(* Logix 5000 project; controller FV vendor 1 type 14 code 217 rev 31.11; software revision 31.00; part 63 of 63 *)
(* tags used below, declared in another part *)
   Alarm_Reset : BOOL;
   CWD : CHECKWORD_FLAGS;
   Default_Check_Time : DINT;
   Item_Faults_Are_Latched : BOOL;
   Item_Simulation_Flag : BOOL;
   One_Second_One_Scan : ALIAS FOR One_Second_1_scan;
   YP_AV1 : PlantItem;   // AV1
   YP_AV1_ALARM : ALARM_DIGITAL;
   YP_AV1_DR : ALIAS FOR RIO_Rack_3:3:O.Data.3;
   YP_AV1_O : ALIAS FOR RIO_Rack_3:1:I.Data.0;
   YP_AV2 : PlantItem;   // AV2
   YP_AV2_ALARM : ALARM_DIGITAL;
   YP_AV2_DR : ALIAS FOR RIO_Rack_3:3:O.Data.5;
   YP_AV2_O : ALIAS FOR RIO_Rack_3:1:I.Data.2;
   YP_AV3 : PlantItem;   // AV3
   YP_AV3_ALARM : ALARM_DIGITAL;
   YP_AV3_DR : ALIAS FOR RIO_Rack_3:3:O.Data.6;
   YP_AV3_O : ALIAS FOR RIO_Rack_3:1:I.Data.4;
   YP_AV4 : PlantItem;   // AV4
   YP_AV4_ALARM : ALARM_DIGITAL;
   YP_AV4_DR : ALIAS FOR RIO_Rack_3:3:O.Data.7;
   YP_AV4_O : ALIAS FOR RIO_Rack_3:1:I.Data.6;
   YP_AV5 : PlantItem;   // AV5
   YP_AV5_ALARM : ALARM_DIGITAL;
   YP_AV5_DR : ALIAS FOR RIO_Rack_3:3:O.Data.8;
   YP_AV5_O : ALIAS FOR RIO_Rack_3:1:I.Data.8;
   YP_AV6 : PlantItem;   // AV6
   YP_AV6_ALARM : ALARM_DIGITAL;
   YP_AV6_DR : ALIAS FOR RIO_Rack_3:3:O.Data.9;
   YP_AV6_O : ALIAS FOR RIO_Rack_3:1:I.Data.10;
   YP_AV7 : PlantItem;   // AV7
   YP_AV7_ALARM : ALARM_DIGITAL;
   YP_AV7_DR : ALIAS FOR RIO_Rack_3:3:O.Data.10;
   YP_AV7_O : ALIAS FOR RIO_Rack_3:1:I.Data.12;
   YP_AV8 : PlantItem;   // AV8
   YP_AV8_ALARM : ALARM_DIGITAL;
   YP_AV8_DR : ALIAS FOR RIO_Rack_3:3:O.Data.11;
   YP_AV8_O : ALIAS FOR RIO_Rack_3:1:I.Data.14;
   YP_B103 : INT[15];   // Original N File From SLC, No Description Available
   YP_B3 : INT[7];   // BINARY
   YP_B30 : INT[37];   // Original N File From SLC, No Description Available
   YP_N40 : INT[9];   // Original N File From SLC, No Description Available
   YP_N50 : INT[15];   // Original N File From SLC, No Description Available
   YP_N55 : INT[244];   // Original N File From SLC, No Description Available
   YP_N7 : INT[56];   // INTEGER
   YP_T4 : TIMER[16];   // TIMER
   YP_YST1_HL : PlantItem;   // YST1_HL
   YP_YST2_HL : PlantItem;   // YST2_HL
(* YP_Common, continued *)

ROUTINE YP_RQD_FLAGS_17   (* ladder *)
   0: [XIC(YP_N40[0].1) ,XIC(YP_N40[1].1) ]OTE(YP_B30[0].1);
   1: [XIC(YP_N40[0].3) ,XIC(YP_N40[0].4) ]XIC(YP_B3[0].10)XIC(YP_B3[0].8)[XIC(YP_B3[0].0) ,XIC(YP_B3[0].2) ,XIC(YP_B3[0].4) ,XIC(YP_B3[0].6) ]OTE(YP_B30[0].4);
   2: [[XIC(YP_N40[0].3) ,XIC(YP_N40[0].4) ,XIC(YP_B103[2].0) ] EQU(YP_N50[5],0) ,EQU(YP_N50[5],1) ]OTE(YP_B30[0].9);
   3: [[XIC(YP_N40[0].3) ,XIC(YP_N40[0].4) ,XIC(YP_B103[2].1) ] EQU(YP_N50[4],0) ,EQU(YP_N50[4],1) ]OTE(YP_B30[0].8);
   4: [[XIC(YP_N40[0].3) ,XIC(YP_N40[0].4) ,XIC(YP_B103[2].0) ,XIC(YP_B103[2].1) ] EQU(YP_N50[0],0) ,EQU(YP_N50[0],1) ]OTE(YP_B30[0].3);
   5: [[XIC(YP_N40[0].3) ,XIC(YP_N40[0].4) ,XIC(YP_B103[2].0) ] EQU(YP_N50[1],0) ,EQU(YP_N50[1],1) ]OTE(YP_B30[0].5);
   6: [[XIC(YP_N40[0].4) ,XIC(YP_B103[2].0) ] EQU(YP_N50[2],0) ,EQU(YP_N50[2],1) ]OTE(YP_B30[0].6);
   7: [[XIC(YP_N40[0].4) ,XIC(YP_B103[2].0) ] EQU(YP_N50[3],0) ,EQU(YP_N50[3],1) ]OTE(YP_B30[0].7);
   8: [XIC(YP_N40[0].7) ,XIC(YP_N40[1].5) ]OTE(YP_B30[0].0);
   9: XIC(YP_N40[0].8)OTE(YP_B30[0].2);
   10: [XIC(YP_N40[2].1) EQU(YP_N50[7],0) ,EQU(YP_N50[7],1) ]OTE(YP_B30[0].11);
   11: [XIC(YP_N40[3].1) EQU(YP_N50[6],0) XIO(YP_N7[38].0) XIO(YP_N7[38].1) ,EQU(YP_N50[6],1) ]OTE(YP_B30[0].10);
   12: [[XIC(YP_N40[0].3) ,XIC(YP_N40[0].4) ] XIC(YP_B3[0].10) XIC(YP_B3[0].8) [XIC(YP_B3[0].0) ,XIC(YP_B3[0].2) ,XIC(YP_B3[0].4) ,XIC(YP_B3[0].6) ] EQU(YP_N50[8],0) ,EQU(YP_N50[8],1) ]OTE(YP_B30[0].12);
   13: [XIC(YP_N40[3].1) XIC(YP_B3[0].12) EQU(YP_N50[9],0) ,EQU(YP_N50[9],1) ]OTE(YP_B30[0].14);
   14: XIC(YP_N40[0].0)MOV(0,YP_N55[2]);
   15: [XIC(YP_N40[0].1) ,XIC(YP_N40[1].1) ]MOV(1,YP_N55[2]);
   16: [XIC(YP_N40[0].2) ,XIC(YP_N40[1].2) ]MOV(2,YP_N55[2]);
   17: XIC(YP_N40[0].3)MOV(3,YP_N55[2]);
   18: XIC(YP_N40[0].4)MOV(4,YP_N55[2]);
   19: XIC(YP_N40[0].5)MOV(5,YP_N55[2]);
   20: XIC(YP_N40[0].6)MOV(6,YP_N55[2]);
   21: [XIC(YP_N40[0].7) ,XIC(YP_N40[1].5) ]MOV(7,YP_N55[2]);
   22: XIC(YP_N40[0].8)MOV(8,YP_N55[2]);
   23: EQU(YP_N55[0],1)MOV(9,YP_N55[2]);
   24: XIC(YP_N40[1].2)MOV(10,YP_N55[2]);
   25: XIC(YP_N40[1].3)MOV(11,YP_N55[2]);
   26: XIC(YP_N40[1].4)MOV(12,YP_N55[2]);
END_ROUTINE

ROUTINE YP_Valves   (* ladder *)
   0: [NEQ(YP_AV1.DriveBits,0) OTE(YP_AV1.CW.[CWD.AUTODRV]) ,[XIC(YP_AV1.CW.[CWD.AUTODRV]) XIO(YP_AV1.CW.[CWD.MANUAL]) ,XIC(YP_AV1.CW.[CWD.MANDRV]) XIC(YP_AV1.CW.[CWD.MANUAL]) ] OTE(YP_AV1.CW.[CWD.OUTPUT]) ,XIC(YP_AV1.CW.[CWD.OUTPUT]) OTE(YP_AV1_DR) ,XIC(S:FS) [OTU(YP_AV1.CW.[CWD.MANUAL]) ,LEQ(YP_AV1.CheckTime,0) MOV(Default_Check_Time,YP_AV1.CheckTime) ] ,[[XIC(YP_AV1_O) XIO(Item_Simulation_Flag) ,XIC(Item_Simulation_Flag) XIC(YP_AV1.CW.[CWD.OUTPUT]) XIO(YP_AV1.CW.[CWD.SIMFAIL]) ] OTE(YP_AV1.CW.[CWD.OPENFB]) ,[XIO(YP_AV1_O) XIO(Item_Simulation_Flag) ,XIC(Item_Simulation_Flag) XIO(YP_AV1.CW.[CWD.OUTPUT]) XIO(YP_AV1.CW.[CWD.SIMFAIL]) ] OTE(YP_AV1.CW.[CWD.CLOSEDFB]) ] ,[XIC(YP_AV1.CW.[CWD.OUTPUT]) XIO(YP_AV1.CW.[CWD.PREVSCAN]) ,XIO(YP_AV1.CW.[CWD.OUTPUT]) XIC(YP_AV1.CW.[CWD.PREVSCAN]) ] CLR(YP_AV1.CheckTimer) ,XIC(One_Second_One_Scan) LES(YP_AV1.CheckTimer,YP_AV1.CheckTime) ADD(YP_AV1.CheckTimer,1,YP_AV1.CheckTimer) ,XIO(YP_AV1.CW.[CWD.FAULT]) OTU(YP_AV1.CW.[CWD.FAULTLOGGED]) ,[GEQ(YP_AV1.CheckTimer,YP_AV1.CheckTime) [XIC(YP_AV1.CW.[CWD.OUTPUT]) [XIO(YP_AV1.CW.[CWD.OPENFB]) ,XIC(YP_AV1.CW.[CWD.CLOSEDFB]) ] ,XIO(YP_AV1.CW.[CWD.OUTPUT]) [XIC(YP_AV1.CW.[CWD.OPENFB]) ,XIO(YP_AV1.CW.[CWD.CLOSEDFB]) ] ] ,XIC(YP_AV1.CW.[CWD.FAULT]) XIC(Item_Faults_Are_Latched) ,XIC(YP_AV1.CW.[CWD.HIGHLIGHT]) ] XIO(YP_AV1.CW.[CWD.CHECKOFF]) XIO(Alarm_Reset) [OTE(YP_AV1.CW.[CWD.FAULT]) ,ALMD(YP_AV1_ALARM,0,0,0,0) ] ,XIC(YP_AV1.CW.[CWD.OUTPUT]) OTE(YP_AV1.CW.[CWD.PREVSCAN]) ];
   1: [NEQ(YP_AV2.DriveBits,0) OTE(YP_AV2.CW.[CWD.AUTODRV]) ,[XIC(YP_AV2.CW.[CWD.AUTODRV]) XIO(YP_AV2.CW.[CWD.MANUAL]) ,XIC(YP_AV2.CW.[CWD.MANDRV]) XIC(YP_AV2.CW.[CWD.MANUAL]) ] OTE(YP_AV2.CW.[CWD.OUTPUT]) ,XIC(YP_AV2.CW.[CWD.OUTPUT]) OTE(YP_AV2_DR) ,XIC(S:FS) [OTU(YP_AV2.CW.[CWD.MANUAL]) ,LEQ(YP_AV2.CheckTime,0) MOV(Default_Check_Time,YP_AV2.CheckTime) ] ,[[XIC(YP_AV2_O) XIO(Item_Simulation_Flag) ,XIC(Item_Simulation_Flag) XIC(YP_AV2.CW.[CWD.OUTPUT]) XIO(YP_AV2.CW.[CWD.SIMFAIL]) ] OTE(YP_AV2.CW.[CWD.OPENFB]) ,[XIO(YP_AV2_O) XIO(Item_Simulation_Flag) ,XIC(Item_Simulation_Flag) XIO(YP_AV2.CW.[CWD.OUTPUT]) XIO(YP_AV2.CW.[CWD.SIMFAIL]) ] OTE(YP_AV2.CW.[CWD.CLOSEDFB]) ] ,[XIC(YP_AV2.CW.[CWD.OUTPUT]) XIO(YP_AV2.CW.[CWD.PREVSCAN]) ,XIO(YP_AV2.CW.[CWD.OUTPUT]) XIC(YP_AV2.CW.[CWD.PREVSCAN]) ] CLR(YP_AV2.CheckTimer) ,XIC(One_Second_One_Scan) LES(YP_AV2.CheckTimer,YP_AV2.CheckTime) ADD(YP_AV2.CheckTimer,1,YP_AV2.CheckTimer) ,XIO(YP_AV2.CW.[CWD.FAULT]) OTU(YP_AV2.CW.[CWD.FAULTLOGGED]) ,[GEQ(YP_AV2.CheckTimer,YP_AV2.CheckTime) [XIC(YP_AV2.CW.[CWD.OUTPUT]) [XIO(YP_AV2.CW.[CWD.OPENFB]) ,XIC(YP_AV2.CW.[CWD.CLOSEDFB]) ] ,XIO(YP_AV2.CW.[CWD.OUTPUT]) [XIC(YP_AV2.CW.[CWD.OPENFB]) ,XIO(YP_AV2.CW.[CWD.CLOSEDFB]) ] ] ,XIC(YP_AV2.CW.[CWD.FAULT]) XIC(Item_Faults_Are_Latched) ,XIC(YP_AV2.CW.[CWD.HIGHLIGHT]) ] XIO(YP_AV2.CW.[CWD.CHECKOFF]) XIO(Alarm_Reset) [OTE(YP_AV2.CW.[CWD.FAULT]) ,ALMD(YP_AV2_ALARM,0,0,0,0) ] ,XIC(YP_AV2.CW.[CWD.OUTPUT]) OTE(YP_AV2.CW.[CWD.PREVSCAN]) ];
   2: [NEQ(YP_AV3.DriveBits,0) OTE(YP_AV3.CW.[CWD.AUTODRV]) ,[XIC(YP_AV3.CW.[CWD.AUTODRV]) XIO(YP_AV3.CW.[CWD.MANUAL]) ,XIC(YP_AV3.CW.[CWD.MANDRV]) XIC(YP_AV3.CW.[CWD.MANUAL]) ] OTE(YP_AV3.CW.[CWD.OUTPUT]) ,XIC(YP_AV3.CW.[CWD.OUTPUT]) OTE(YP_AV3_DR) ,XIC(S:FS) [OTU(YP_AV3.CW.[CWD.MANUAL]) ,LEQ(YP_AV3.CheckTime,0) MOV(Default_Check_Time,YP_AV3.CheckTime) ] ,[[XIC(YP_AV3_O) XIO(Item_Simulation_Flag) ,XIC(Item_Simulation_Flag) XIC(YP_AV3.CW.[CWD.OUTPUT]) XIO(YP_AV3.CW.[CWD.SIMFAIL]) ] OTE(YP_AV3.CW.[CWD.OPENFB]) ,[XIO(YP_AV3_O) XIO(Item_Simulation_Flag) ,XIC(Item_Simulation_Flag) XIO(YP_AV3.CW.[CWD.OUTPUT]) XIO(YP_AV3.CW.[CWD.SIMFAIL]) ] OTE(YP_AV3.CW.[CWD.CLOSEDFB]) ] ,[XIC(YP_AV3.CW.[CWD.OUTPUT]) XIO(YP_AV3.CW.[CWD.PREVSCAN]) ,XIO(YP_AV3.CW.[CWD.OUTPUT]) XIC(YP_AV3.CW.[CWD.PREVSCAN]) ] CLR(YP_AV3.CheckTimer) ,XIC(One_Second_One_Scan) LES(YP_AV3.CheckTimer,YP_AV3.CheckTime) ADD(YP_AV3.CheckTimer,1,YP_AV3.CheckTimer) ,XIO(YP_AV3.CW.[CWD.FAULT]) OTU(YP_AV3.CW.[CWD.FAULTLOGGED]) ,[GEQ(YP_AV3.CheckTimer,YP_AV3.CheckTime) [XIC(YP_AV3.CW.[CWD.OUTPUT]) [XIO(YP_AV3.CW.[CWD.OPENFB]) ,XIC(YP_AV3.CW.[CWD.CLOSEDFB]) ] ,XIO(YP_AV3.CW.[CWD.OUTPUT]) [XIC(YP_AV3.CW.[CWD.OPENFB]) ,XIO(YP_AV3.CW.[CWD.CLOSEDFB]) ] ] ,XIC(YP_AV3.CW.[CWD.FAULT]) XIC(Item_Faults_Are_Latched) ,XIC(YP_AV3.CW.[CWD.HIGHLIGHT]) ] XIO(YP_AV3.CW.[CWD.CHECKOFF]) XIO(Alarm_Reset) [OTE(YP_AV3.CW.[CWD.FAULT]) ,ALMD(YP_AV3_ALARM,0,0,0,0) ] ,XIC(YP_AV3.CW.[CWD.OUTPUT]) OTE(YP_AV3.CW.[CWD.PREVSCAN]) ];
   3: [NEQ(YP_AV4.DriveBits,0) OTE(YP_AV4.CW.[CWD.AUTODRV]) ,[XIC(YP_AV4.CW.[CWD.AUTODRV]) XIO(YP_AV4.CW.[CWD.MANUAL]) ,XIC(YP_AV4.CW.[CWD.MANDRV]) XIC(YP_AV4.CW.[CWD.MANUAL]) ] OTE(YP_AV4.CW.[CWD.OUTPUT]) ,XIC(YP_AV4.CW.[CWD.OUTPUT]) OTE(YP_AV4_DR) ,XIC(S:FS) [OTU(YP_AV4.CW.[CWD.MANUAL]) ,LEQ(YP_AV4.CheckTime,0) MOV(Default_Check_Time,YP_AV4.CheckTime) ] ,[[XIC(YP_AV4_O) XIO(Item_Simulation_Flag) ,XIC(Item_Simulation_Flag) XIC(YP_AV4.CW.[CWD.OUTPUT]) XIO(YP_AV4.CW.[CWD.SIMFAIL]) ] OTE(YP_AV4.CW.[CWD.OPENFB]) ,[XIO(YP_AV4_O) XIO(Item_Simulation_Flag) ,XIC(Item_Simulation_Flag) XIO(YP_AV4.CW.[CWD.OUTPUT]) XIO(YP_AV4.CW.[CWD.SIMFAIL]) ] OTE(YP_AV4.CW.[CWD.CLOSEDFB]) ] ,[XIC(YP_AV4.CW.[CWD.OUTPUT]) XIO(YP_AV4.CW.[CWD.PREVSCAN]) ,XIO(YP_AV4.CW.[CWD.OUTPUT]) XIC(YP_AV4.CW.[CWD.PREVSCAN]) ] CLR(YP_AV4.CheckTimer) ,XIC(One_Second_One_Scan) LES(YP_AV4.CheckTimer,YP_AV4.CheckTime) ADD(YP_AV4.CheckTimer,1,YP_AV4.CheckTimer) ,XIO(YP_AV4.CW.[CWD.FAULT]) OTU(YP_AV4.CW.[CWD.FAULTLOGGED]) ,[GEQ(YP_AV4.CheckTimer,YP_AV4.CheckTime) [XIC(YP_AV4.CW.[CWD.OUTPUT]) [XIO(YP_AV4.CW.[CWD.OPENFB]) ,XIC(YP_AV4.CW.[CWD.CLOSEDFB]) ] ,XIO(YP_AV4.CW.[CWD.OUTPUT]) [XIC(YP_AV4.CW.[CWD.OPENFB]) ,XIO(YP_AV4.CW.[CWD.CLOSEDFB]) ] ] ,XIC(YP_AV4.CW.[CWD.FAULT]) XIC(Item_Faults_Are_Latched) ,XIC(YP_AV4.CW.[CWD.HIGHLIGHT]) ] XIO(YP_AV4.CW.[CWD.CHECKOFF]) XIO(Alarm_Reset) [OTE(YP_AV4.CW.[CWD.FAULT]) ,ALMD(YP_AV4_ALARM,0,0,0,0) ] ,XIC(YP_AV4.CW.[CWD.OUTPUT]) OTE(YP_AV4.CW.[CWD.PREVSCAN]) ];
   4: [NEQ(YP_AV5.DriveBits,0) OTE(YP_AV5.CW.[CWD.AUTODRV]) ,[XIC(YP_AV5.CW.[CWD.AUTODRV]) XIO(YP_AV5.CW.[CWD.MANUAL]) ,XIC(YP_AV5.CW.[CWD.MANDRV]) XIC(YP_AV5.CW.[CWD.MANUAL]) ] OTE(YP_AV5.CW.[CWD.OUTPUT]) ,XIC(YP_AV5.CW.[CWD.OUTPUT]) OTE(YP_AV5_DR) ,XIC(S:FS) [OTU(YP_AV5.CW.[CWD.MANUAL]) ,LEQ(YP_AV5.CheckTime,0) MOV(Default_Check_Time,YP_AV5.CheckTime) ] ,[[XIC(YP_AV5_O) XIO(Item_Simulation_Flag) ,XIC(Item_Simulation_Flag) XIC(YP_AV5.CW.[CWD.OUTPUT]) XIO(YP_AV5.CW.[CWD.SIMFAIL]) ] OTE(YP_AV5.CW.[CWD.OPENFB]) ,[XIO(YP_AV5_O) XIO(Item_Simulation_Flag) ,XIC(Item_Simulation_Flag) XIO(YP_AV5.CW.[CWD.OUTPUT]) XIO(YP_AV5.CW.[CWD.SIMFAIL]) ] OTE(YP_AV5.CW.[CWD.CLOSEDFB]) ] ,[XIC(YP_AV5.CW.[CWD.OUTPUT]) XIO(YP_AV5.CW.[CWD.PREVSCAN]) ,XIO(YP_AV5.CW.[CWD.OUTPUT]) XIC(YP_AV5.CW.[CWD.PREVSCAN]) ] CLR(YP_AV5.CheckTimer) ,XIC(One_Second_One_Scan) LES(YP_AV5.CheckTimer,YP_AV5.CheckTime) ADD(YP_AV5.CheckTimer,1,YP_AV5.CheckTimer) ,XIO(YP_AV5.CW.[CWD.FAULT]) OTU(YP_AV5.CW.[CWD.FAULTLOGGED]) ,[GEQ(YP_AV5.CheckTimer,YP_AV5.CheckTime) [XIC(YP_AV5.CW.[CWD.OUTPUT]) [XIO(YP_AV5.CW.[CWD.OPENFB]) ,XIC(YP_AV5.CW.[CWD.CLOSEDFB]) ] ,XIO(YP_AV5.CW.[CWD.OUTPUT]) [XIC(YP_AV5.CW.[CWD.OPENFB]) ,XIO(YP_AV5.CW.[CWD.CLOSEDFB]) ] ] ,XIC(YP_AV5.CW.[CWD.FAULT]) XIC(Item_Faults_Are_Latched) ,XIC(YP_AV5.CW.[CWD.HIGHLIGHT]) ] XIO(YP_AV5.CW.[CWD.CHECKOFF]) XIO(Alarm_Reset) [OTE(YP_AV5.CW.[CWD.FAULT]) ,ALMD(YP_AV5_ALARM,0,0,0,0) ] ,XIC(YP_AV5.CW.[CWD.OUTPUT]) OTE(YP_AV5.CW.[CWD.PREVSCAN]) ];
   5: [NEQ(YP_AV6.DriveBits,0) OTE(YP_AV6.CW.[CWD.AUTODRV]) ,[XIC(YP_AV6.CW.[CWD.AUTODRV]) XIO(YP_AV6.CW.[CWD.MANUAL]) ,XIC(YP_AV6.CW.[CWD.MANDRV]) XIC(YP_AV6.CW.[CWD.MANUAL]) ] OTE(YP_AV6.CW.[CWD.OUTPUT]) ,XIC(YP_AV6.CW.[CWD.OUTPUT]) OTE(YP_AV6_DR) ,XIC(S:FS) [OTU(YP_AV6.CW.[CWD.MANUAL]) ,LEQ(YP_AV6.CheckTime,0) MOV(Default_Check_Time,YP_AV6.CheckTime) ] ,[[XIC(YP_AV6_O) XIO(Item_Simulation_Flag) ,XIC(Item_Simulation_Flag) XIC(YP_AV6.CW.[CWD.OUTPUT]) XIO(YP_AV6.CW.[CWD.SIMFAIL]) ] OTE(YP_AV6.CW.[CWD.OPENFB]) ,[XIO(YP_AV6_O) XIO(Item_Simulation_Flag) ,XIC(Item_Simulation_Flag) XIO(YP_AV6.CW.[CWD.OUTPUT]) XIO(YP_AV6.CW.[CWD.SIMFAIL]) ] OTE(YP_AV6.CW.[CWD.CLOSEDFB]) ] ,[XIC(YP_AV6.CW.[CWD.OUTPUT]) XIO(YP_AV6.CW.[CWD.PREVSCAN]) ,XIO(YP_AV6.CW.[CWD.OUTPUT]) XIC(YP_AV6.CW.[CWD.PREVSCAN]) ] CLR(YP_AV6.CheckTimer) ,XIC(One_Second_One_Scan) LES(YP_AV6.CheckTimer,YP_AV6.CheckTime) ADD(YP_AV6.CheckTimer,1,YP_AV6.CheckTimer) ,XIO(YP_AV6.CW.[CWD.FAULT]) OTU(YP_AV6.CW.[CWD.FAULTLOGGED]) ,[GEQ(YP_AV6.CheckTimer,YP_AV6.CheckTime) [XIC(YP_AV6.CW.[CWD.OUTPUT]) [XIO(YP_AV6.CW.[CWD.OPENFB]) ,XIC(YP_AV6.CW.[CWD.CLOSEDFB]) ] ,XIO(YP_AV6.CW.[CWD.OUTPUT]) [XIC(YP_AV6.CW.[CWD.OPENFB]) ,XIO(YP_AV6.CW.[CWD.CLOSEDFB]) ] ] ,XIC(YP_AV6.CW.[CWD.FAULT]) XIC(Item_Faults_Are_Latched) ,XIC(YP_AV6.CW.[CWD.HIGHLIGHT]) ] XIO(YP_AV6.CW.[CWD.CHECKOFF]) XIO(Alarm_Reset) [OTE(YP_AV6.CW.[CWD.FAULT]) ,ALMD(YP_AV6_ALARM,0,0,0,0) ] ,XIC(YP_AV6.CW.[CWD.OUTPUT]) OTE(YP_AV6.CW.[CWD.PREVSCAN]) ];
   6: [NEQ(YP_AV7.DriveBits,0) OTE(YP_AV7.CW.[CWD.AUTODRV]) ,[XIC(YP_AV7.CW.[CWD.AUTODRV]) XIO(YP_AV7.CW.[CWD.MANUAL]) ,XIC(YP_AV7.CW.[CWD.MANDRV]) XIC(YP_AV7.CW.[CWD.MANUAL]) ] OTE(YP_AV7.CW.[CWD.OUTPUT]) ,XIC(YP_AV7.CW.[CWD.OUTPUT]) OTE(YP_AV7_DR) ,XIC(S:FS) [OTU(YP_AV7.CW.[CWD.MANUAL]) ,LEQ(YP_AV7.CheckTime,0) MOV(Default_Check_Time,YP_AV7.CheckTime) ] ,[[XIC(YP_AV7_O) XIO(Item_Simulation_Flag) ,XIC(Item_Simulation_Flag) XIC(YP_AV7.CW.[CWD.OUTPUT]) XIO(YP_AV7.CW.[CWD.SIMFAIL]) ] OTE(YP_AV7.CW.[CWD.OPENFB]) ,[XIO(YP_AV7_O) XIO(Item_Simulation_Flag) ,XIC(Item_Simulation_Flag) XIO(YP_AV7.CW.[CWD.OUTPUT]) XIO(YP_AV7.CW.[CWD.SIMFAIL]) ] OTE(YP_AV7.CW.[CWD.CLOSEDFB]) ] ,[XIC(YP_AV7.CW.[CWD.OUTPUT]) XIO(YP_AV7.CW.[CWD.PREVSCAN]) ,XIO(YP_AV7.CW.[CWD.OUTPUT]) XIC(YP_AV7.CW.[CWD.PREVSCAN]) ] CLR(YP_AV7.CheckTimer) ,XIC(One_Second_One_Scan) LES(YP_AV7.CheckTimer,YP_AV7.CheckTime) ADD(YP_AV7.CheckTimer,1,YP_AV7.CheckTimer) ,XIO(YP_AV7.CW.[CWD.FAULT]) OTU(YP_AV7.CW.[CWD.FAULTLOGGED]) ,[GEQ(YP_AV7.CheckTimer,YP_AV7.CheckTime) [XIC(YP_AV7.CW.[CWD.OUTPUT]) [XIO(YP_AV7.CW.[CWD.OPENFB]) ,XIC(YP_AV7.CW.[CWD.CLOSEDFB]) ] ,XIO(YP_AV7.CW.[CWD.OUTPUT]) [XIC(YP_AV7.CW.[CWD.OPENFB]) ,XIO(YP_AV7.CW.[CWD.CLOSEDFB]) ] ] ,XIC(YP_AV7.CW.[CWD.FAULT]) XIC(Item_Faults_Are_Latched) ,XIC(YP_AV7.CW.[CWD.HIGHLIGHT]) ] XIO(YP_AV7.CW.[CWD.CHECKOFF]) XIO(Alarm_Reset) [OTE(YP_AV7.CW.[CWD.FAULT]) ,ALMD(YP_AV7_ALARM,0,0,0,0) ] ,XIC(YP_AV7.CW.[CWD.OUTPUT]) OTE(YP_AV7.CW.[CWD.PREVSCAN]) ];
   7: [NEQ(YP_AV8.DriveBits,0) OTE(YP_AV8.CW.[CWD.AUTODRV]) ,[XIC(YP_AV8.CW.[CWD.AUTODRV]) XIO(YP_AV8.CW.[CWD.MANUAL]) ,XIC(YP_AV8.CW.[CWD.MANDRV]) XIC(YP_AV8.CW.[CWD.MANUAL]) ] OTE(YP_AV8.CW.[CWD.OUTPUT]) ,XIC(YP_AV8.CW.[CWD.OUTPUT]) OTE(YP_AV8_DR) ,XIC(S:FS) [OTU(YP_AV8.CW.[CWD.MANUAL]) ,LEQ(YP_AV8.CheckTime,0) MOV(Default_Check_Time,YP_AV8.CheckTime) ] ,[[XIC(YP_AV8_O) XIO(Item_Simulation_Flag) ,XIC(Item_Simulation_Flag) XIC(YP_AV8.CW.[CWD.OUTPUT]) XIO(YP_AV8.CW.[CWD.SIMFAIL]) ] OTE(YP_AV8.CW.[CWD.OPENFB]) ,[XIO(YP_AV8_O) XIO(Item_Simulation_Flag) ,XIC(Item_Simulation_Flag) XIO(YP_AV8.CW.[CWD.OUTPUT]) XIO(YP_AV8.CW.[CWD.SIMFAIL]) ] OTE(YP_AV8.CW.[CWD.CLOSEDFB]) ] ,[XIC(YP_AV8.CW.[CWD.OUTPUT]) XIO(YP_AV8.CW.[CWD.PREVSCAN]) ,XIO(YP_AV8.CW.[CWD.OUTPUT]) XIC(YP_AV8.CW.[CWD.PREVSCAN]) ] CLR(YP_AV8.CheckTimer) ,XIC(One_Second_One_Scan) LES(YP_AV8.CheckTimer,YP_AV8.CheckTime) ADD(YP_AV8.CheckTimer,1,YP_AV8.CheckTimer) ,XIO(YP_AV8.CW.[CWD.FAULT]) OTU(YP_AV8.CW.[CWD.FAULTLOGGED]) ,[GEQ(YP_AV8.CheckTimer,YP_AV8.CheckTime) [XIC(YP_AV8.CW.[CWD.OUTPUT]) [XIO(YP_AV8.CW.[CWD.OPENFB]) ,XIC(YP_AV8.CW.[CWD.CLOSEDFB]) ] ,XIO(YP_AV8.CW.[CWD.OUTPUT]) [XIC(YP_AV8.CW.[CWD.OPENFB]) ,XIO(YP_AV8.CW.[CWD.CLOSEDFB]) ] ] ,XIC(YP_AV8.CW.[CWD.FAULT]) XIC(Item_Faults_Are_Latched) ,XIC(YP_AV8.CW.[CWD.HIGHLIGHT]) ] XIO(YP_AV8.CW.[CWD.CHECKOFF]) XIO(Alarm_Reset) [OTE(YP_AV8.CW.[CWD.FAULT]) ,ALMD(YP_AV8_ALARM,0,0,0,0) ] ,XIC(YP_AV8.CW.[CWD.OUTPUT]) OTE(YP_AV8.CW.[CWD.PREVSCAN]) ];
END_ROUTINE

ROUTINE YP_YSTS_HL_18   (* ladder *)
   0: XIO(YP_YST1_HL.CW.[CWD.INPUTSTATUS])[TON(YP_T4[4],?,?) ,XIC(YP_T4[4].DN) OTL(YP_N7[40].0) ];
   1: XIC(YP_YST1_HL.CW.[CWD.INPUTSTATUS])[TON(YP_T4[5],?,?) ,XIC(YP_T4[5].DN) OTU(YP_N7[40].0) ];
   2: XIO(YP_YST2_HL.CW.[CWD.INPUTSTATUS])[TON(YP_T4[6],?,?) ,XIC(YP_T4[6].DN) OTL(YP_N7[40].1) ];
   3: XIC(YP_YST2_HL.CW.[CWD.INPUTSTATUS])[TON(YP_T4[7],?,?) ,XIC(YP_T4[7].DN) OTU(YP_N7[40].1) ];
END_ROUTINE
END_PROGRAM
